   // TANK_CONTROL_6S.GTT_OUT_DATA.GTT_DemandsCompleted[2] := False;
   // TANK_CONTROL_6S.GTT_OUT_DATA.GTT_DemandsCompleted[1] := False;
   // TANK_CONTROL_6S.PVVX_OUT_DATA.PVVB_Alarms[14] := False;
   // TANK_CONTROL_6S.PVVX_OUT_DATA.PVVB_Alarms[13] := False;
   // TANK_CONTROL_6S.PVVX_OUT_DATA.PVVB_Alarms[12] := False;
   // TANK_CONTROL_6S.PVVX_OUT_DATA.PVVB_Alarms[11] := False;
   // TANK_CONTROL_6S.PVVX_OUT_DATA.PVVB_Alarms[10] := False;
   // TANK_CONTROL_6S.PVVX_OUT_DATA.PVVB_Alarms[9] := False;
   // TANK_CONTROL_6S.PVVX_OUT_DATA.PVVB_Alarms[8] := False;
   // TANK_CONTROL_6S.PVVX_OUT_DATA.PVVB_Alarms[7] := False;
   // TANK_CONTROL_6S.PVVX_OUT_DATA.PVVB_Alarms[6] := False;
   // TANK_CONTROL_6S.PVVX_OUT_DATA.PVVB_Alarms[5] := False;
   // TANK_CONTROL_6S.PVVX_OUT_DATA.PVVB_Alarms[4] := False;
   // TANK_CONTROL_6S.PVVX_OUT_DATA.PVVB_Alarms[3] := False;
   // TANK_CONTROL_6S.PVVX_OUT_DATA.PVVB_Alarms[2] := False;
   // TANK_CONTROL_6S.PVVX_OUT_DATA.PVVB_Alarms[1] := False;
   // TANK_CONTROL_6S.PVVX_OUT_DATA.PVVB_DemandsCompleted[14] := False;
   // TANK_CONTROL_6S.PVVX_OUT_DATA.PVVB_DemandsCompleted[13] := False;
   // TANK_CONTROL_6S.PVVX_OUT_DATA.PVVB_DemandsCompleted[12] := False;
   // TANK_CONTROL_6S.PVVX_OUT_DATA.PVVB_DemandsCompleted[11] := False;
   // TANK_CONTROL_6S.PVVX_OUT_DATA.PVVB_DemandsCompleted[10] := False;
   // TANK_CONTROL_6S.PVVX_OUT_DATA.PVVB_DemandsCompleted[9] := False;
   // TANK_CONTROL_6S.PVVX_OUT_DATA.PVVB_DemandsCompleted[8] := False;
   // TANK_CONTROL_6S.PVVX_OUT_DATA.PVVB_DemandsCompleted[7] := False;
   // TANK_CONTROL_6S.PVVX_OUT_DATA.PVVB_DemandsCompleted[6] := False;
   // TANK_CONTROL_6S.PVVX_OUT_DATA.PVVB_DemandsCompleted[5] := False;
   // TANK_CONTROL_6S.PVVX_OUT_DATA.PVVB_DemandsCompleted[4] := False;
   // TANK_CONTROL_6S.PVVX_OUT_DATA.PVVB_DemandsCompleted[3] := False;
   // TANK_CONTROL_6S.PVVX_OUT_DATA.PVVB_DemandsCompleted[2] := False;
   // TANK_CONTROL_6S.PVVX_OUT_DATA.PVVB_DemandsCompleted[1] := False;
   // TANK_CONTROL_6S.PVVX_OUT_DATA.PVVA_Alarms[14] := False;
   // TANK_CONTROL_6S.PVVX_OUT_DATA.PVVA_Alarms[13] := False;
   // TANK_CONTROL_6S.PVVX_OUT_DATA.PVVA_Alarms[12] := False;
   // TANK_CONTROL_6S.PVVX_OUT_DATA.PVVA_Alarms[11] := False;
   // TANK_CONTROL_6S.PVVX_OUT_DATA.PVVA_Alarms[10] := False;
   // TANK_CONTROL_6S.PVVX_OUT_DATA.PVVA_Alarms[9] := False;
   // TANK_CONTROL_6S.PVVX_OUT_DATA.PVVA_Alarms[8] := False;
   // TANK_CONTROL_6S.PVVX_OUT_DATA.PVVA_Alarms[7] := False;
   // TANK_CONTROL_6S.PVVX_OUT_DATA.PVVA_Alarms[6] := False;
   // TANK_CONTROL_6S.PVVX_OUT_DATA.PVVA_Alarms[5] := False;
   // TANK_CONTROL_6S.PVVX_OUT_DATA.PVVA_Alarms[4] := False;
   // TANK_CONTROL_6S.PVVX_OUT_DATA.PVVA_Alarms[3] := False;
   // TANK_CONTROL_1P.DWELL_TIMER.IN := False;
   // TANK_CONTROL_1P.MONITOR_TIMER.IN := False;
   // TANK_CONTROL_1P.ReOx_InitialTargetpHLevelAchieved := False;
   // TANK_CONTROL_6S.PVVX_OUT_DATA.PVVA_Alarms[2] := False;
   // TANK_CONTROL_6S.PVVX_OUT_DATA.PVVA_Alarms[1] := False;
   // TANK_CONTROL_6S.PVVX_OUT_DATA.PVVA_DemandsCompleted[14] := False;
   // TANK_CONTROL_6S.PVVX_OUT_DATA.PVVA_DemandsCompleted[13] := False;
   // TANK_CONTROL_6S.PVVX_OUT_DATA.PVVA_DemandsCompleted[12] := False;
   // TANK_CONTROL_6S.PVVX_OUT_DATA.PVVA_DemandsCompleted[11] := False;
   // TANK_CONTROL_6S.PVVX_OUT_DATA.PVVA_DemandsCompleted[10] := False;
   // TANK_CONTROL_6S.PVVX_OUT_DATA.PVVA_DemandsCompleted[9] := False;
   // TANK_CONTROL_6S.PVVX_OUT_DATA.PVVA_DemandsCompleted[8] := False;
   // TANK_CONTROL_6S.PVVX_OUT_DATA.PVVA_DemandsCompleted[7] := False;
   // TANK_CONTROL_6S.PVVX_OUT_DATA.PVVA_DemandsCompleted[6] := False;
   // TANK_CONTROL_6S.PVVX_OUT_DATA.PVVA_DemandsCompleted[5] := False;
   // TANK_CONTROL_6S.PVVX_OUT_DATA.PVVA_DemandsCompleted[4] := False;
   // TANK_CONTROL_6S.PVVX_OUT_DATA.PVVA_DemandsCompleted[3] := False;
   // TANK_CONTROL_6S.PVVX_OUT_DATA.PVVA_DemandsCompleted[2] := False;
   // TANK_CONTROL_6S.PVVX_OUT_DATA.PVVA_DemandsCompleted[1] := False;
   // TANK_CONTROL_1P.TankIPData.TANK_GROUP_SPARE_DI_5 := False;
   // TANK_CONTROL_1P.TankIPData.TANK_GROUP_SPARE_DI_6 := False;
   // TANK_CONTROL_1P.TankIPData.TANK_GROUP_SPARE_DI_7 := False;
   // TANK_CONTROL_1P.TankIPData.GTT_ISOL_VALVE_OPEN := False;
   // TANK_CONTROL_1P.TankIPData.GTT_ISOL_VALVE_CLSD := False;
   // TANK_CONTROL_1P.TankIPData.BWT_LEVEL_HIHI := False;
   // TANK_CONTROL_1P.TankIPData.TANK_ALARM := False;
   // TANK_CONTROL_1P.TankIPData.SPARE_DI_7 := False;
   // TANK_CONTROL_1S.TankIPData.TANKS_PRESS_HIHI := False;
   // TANK_CONTROL_1S.TankIPData.TANK_GROUP_SPARE_DI_2 := False;
   // TANK_CONTROL_1S.TankIPData.TANK_GROUP_SPARE_DI_3 := False;
   // TANK_CONTROL_1S.TankIPData.TANK_GROUP_SPARE_DI_4 := False;
   // TANK_CONTROL_1S.TankIPData.TANK_GROUP_SPARE_DI_5 := False;
   // TANK_CONTROL_1S.TankIPData.TANK_GROUP_SPARE_DI_6 := False;
   // TANK_CONTROL_1S.TankIPData.TANK_GROUP_SPARE_DI_7 := False;
   // TANK_CONTROL_1S.TankIPData.GTT_ISOL_VALVE_OPEN := False;
   // TANK_CONTROL_6P.GTT_OUT_DATA.GTT_Alarms[14] := False;
   // TANK_CONTROL_6P.GTT_OUT_DATA.GTT_Alarms[13] := False;
   // TANK_CONTROL_6P.GTT_OUT_DATA.GTT_Alarms[12] := False;
   // TANK_CONTROL_6P.GTT_OUT_DATA.GTT_Alarms[11] := False;
   // TANK_CONTROL_6P.GTT_OUT_DATA.GTT_Alarms[10] := False;
   // TANK_CONTROL_6P.GTT_OUT_DATA.GTT_Alarms[9] := False;
   // TANK_CONTROL_6P.GTT_OUT_DATA.GTT_Alarms[8] := False;
   // TANK_CONTROL_6P.GTT_OUT_DATA.GTT_Alarms[7] := False;
   // TANK_CONTROL_6P.GTT_OUT_DATA.GTT_Alarms[6] := False;
   // TANK_CONTROL_6P.GTT_OUT_DATA.GTT_Alarms[5] := False;
   // TANK_CONTROL_6P.GTT_OUT_DATA.GTT_Alarms[4] := False;
   // TANK_CONTROL_6P.GTT_OUT_DATA.GTT_Alarms[3] := False;
   // TANK_CONTROL_6P.GTT_OUT_DATA.GTT_Alarms[2] := False;
   // TANK_CONTROL_6P.GTT_OUT_DATA.GTT_Alarms[1] := False;
   // TANK_CONTROL_6P.GTT_OUT_DATA.GTT_DemandsCompleted[14] := False;
   // TANK_CONTROL_6P.GTT_OUT_DATA.GTT_DemandsCompleted[13] := False;
   // TANK_CONTROL_6P.GTT_OUT_DATA.GTT_DemandsCompleted[12] := False;
   // TANK_CONTROL_6P.GTT_OUT_DATA.GTT_DemandsCompleted[11] := False;
   // TANK_CONTROL_6P.GTT_OUT_DATA.GTT_DemandsCompleted[10] := False;
   // TANK_CONTROL_6P.GTT_OUT_DATA.GTT_DemandsCompleted[9] := False;
   // TANK_CONTROL_6P.GTT_OUT_DATA.GTT_DemandsCompleted[8] := False;
   // TANK_CONTROL_6P.GTT_OUT_DATA.GTT_DemandsCompleted[7] := False;
   // TANK_CONTROL_6P.GTT_OUT_DATA.GTT_DemandsCompleted[6] := False;
   // TANK_CONTROL_6P.GTT_OUT_DATA.GTT_DemandsCompleted[5] := False;
   // TANK_CONTROL_6P.GTT_OUT_DATA.GTT_DemandsCompleted[4] := False;
   // TANK_CONTROL_6P.GTT_OUT_DATA.GTT_DemandsCompleted[3] := False;
   // TANK_CONTROL_6P.GTT_OUT_DATA.GTT_DemandsCompleted[2] := False;
   // TANK_CONTROL_6P.GTT_OUT_DATA.GTT_DemandsCompleted[1] := False;
   // TANK_CONTROL_6P.PVVX_OUT_DATA.PVVB_Alarms[14] := False;
   // TANK_CONTROL_6P.PVVX_OUT_DATA.PVVB_Alarms[13] := False;
   // TANK_CONTROL_6P.PVVX_OUT_DATA.PVVB_Alarms[12] := False;
   // TANK_CONTROL_6P.PVVX_OUT_DATA.PVVB_Alarms[11] := False;
   // TANK_CONTROL_6P.PVVX_OUT_DATA.PVVB_Alarms[10] := False;
   // TANK_CONTROL_6P.PVVX_OUT_DATA.PVVB_Alarms[9] := False;
   // TANK_CONTROL_6P.PVVX_OUT_DATA.PVVB_Alarms[8] := False;
   // TANK_CONTROL_6P.PVVX_OUT_DATA.PVVB_Alarms[7] := False;
   // TANK_CONTROL_6P.PVVX_OUT_DATA.PVVB_Alarms[6] := False;
   // TANK_CONTROL_6P.PVVX_OUT_DATA.PVVB_Alarms[5] := False;
   // TANK_CONTROL_6P.PVVX_OUT_DATA.PVVB_Alarms[4] := False;
   // TANK_CONTROL_6P.PVVX_OUT_DATA.PVVB_Alarms[3] := False;
   // TANK_CONTROL_6P.PVVX_OUT_DATA.PVVB_Alarms[2] := False;
   // TANK_CONTROL_6P.PVVX_OUT_DATA.PVVB_Alarms[1] := False;
   // TANK_CONTROL_6P.PVVX_OUT_DATA.PVVB_DemandsCompleted[14] := False;
   // TANK_CONTROL_6P.PVVX_OUT_DATA.PVVB_DemandsCompleted[13] := False;
   // TANK_CONTROL_6P.PVVX_OUT_DATA.PVVB_DemandsCompleted[12] := False;
   // TANK_CONTROL_6P.PVVX_OUT_DATA.PVVB_DemandsCompleted[11] := False;
   // TANK_CONTROL_6P.PVVX_OUT_DATA.PVVB_DemandsCompleted[10] := False;
   // TANK_CONTROL_6P.PVVX_OUT_DATA.PVVB_DemandsCompleted[9] := False;
   // TANK_CONTROL_6P.PVVX_OUT_DATA.PVVB_DemandsCompleted[8] := False;
   // TANK_CONTROL_6P.PVVX_OUT_DATA.PVVB_DemandsCompleted[7] := False;
   // TANK_CONTROL_6P.PVVX_OUT_DATA.PVVB_DemandsCompleted[6] := False;
   // TANK_CONTROL_6P.PVVX_OUT_DATA.PVVB_DemandsCompleted[5] := False;
   // TANK_CONTROL_1S.DWELL_TIMER.IN := False;
   // TANK_CONTROL_1S.MONITOR_TIMER.IN := False;
   // TANK_CONTROL_1S.ReOx_InitialTargetpHLevelAchieved := False;
   // TANK_CONTROL_6P.PVVX_OUT_DATA.PVVB_DemandsCompleted[4] := False;
   // TANK_CONTROL_6P.PVVX_OUT_DATA.PVVB_DemandsCompleted[3] := False;
   // TANK_CONTROL_6P.PVVX_OUT_DATA.PVVB_DemandsCompleted[2] := False;
   // TANK_CONTROL_6P.PVVX_OUT_DATA.PVVB_DemandsCompleted[1] := False;
   // TANK_CONTROL_6P.PVVX_OUT_DATA.PVVA_Alarms[14] := False;
   // TANK_CONTROL_6P.PVVX_OUT_DATA.PVVA_Alarms[13] := False;
   // TANK_CONTROL_6P.PVVX_OUT_DATA.PVVA_Alarms[12] := False;
   // TANK_CONTROL_6P.PVVX_OUT_DATA.PVVA_Alarms[11] := False;
   // TANK_CONTROL_6P.PVVX_OUT_DATA.PVVA_Alarms[10] := False;
   // TANK_CONTROL_6P.PVVX_OUT_DATA.PVVA_Alarms[9] := False;
   // TANK_CONTROL_6P.PVVX_OUT_DATA.PVVA_Alarms[8] := False;
   // TANK_CONTROL_6P.PVVX_OUT_DATA.PVVA_Alarms[7] := False;
   // TANK_CONTROL_6P.PVVX_OUT_DATA.PVVA_Alarms[6] := False;
   // TANK_CONTROL_6P.PVVX_OUT_DATA.PVVA_Alarms[5] := False;
   // TANK_CONTROL_6P.PVVX_OUT_DATA.PVVA_Alarms[4] := False;
   // TANK_CONTROL_6P.PVVX_OUT_DATA.PVVA_Alarms[3] := False;
   // TANK_CONTROL_6P.PVVX_OUT_DATA.PVVA_Alarms[2] := False;
   // TANK_CONTROL_6P.PVVX_OUT_DATA.PVVA_Alarms[1] := False;
   // TANK_CONTROL_6P.PVVX_OUT_DATA.PVVA_DemandsCompleted[14] := False;
   // TANK_CONTROL_6P.PVVX_OUT_DATA.PVVA_DemandsCompleted[13] := False;
   // TANK_CONTROL_6P.PVVX_OUT_DATA.PVVA_DemandsCompleted[12] := False;
   // TANK_CONTROL_6P.PVVX_OUT_DATA.PVVA_DemandsCompleted[11] := False;
   // TANK_CONTROL_6P.PVVX_OUT_DATA.PVVA_DemandsCompleted[10] := False;
   // TANK_CONTROL_6P.PVVX_OUT_DATA.PVVA_DemandsCompleted[9] := False;
   // TANK_CONTROL_6P.PVVX_OUT_DATA.PVVA_DemandsCompleted[8] := False;
   // TANK_CONTROL_6P.PVVX_OUT_DATA.PVVA_DemandsCompleted[7] := False;
   // TANK_CONTROL_6P.PVVX_OUT_DATA.PVVA_DemandsCompleted[6] := False;
   // TANK_CONTROL_6P.PVVX_OUT_DATA.PVVA_DemandsCompleted[5] := False;
   // TANK_CONTROL_6P.PVVX_OUT_DATA.PVVA_DemandsCompleted[4] := False;
   // TANK_CONTROL_6P.PVVX_OUT_DATA.PVVA_DemandsCompleted[3] := False;
   // TANK_CONTROL_6P.PVVX_OUT_DATA.PVVA_DemandsCompleted[2] := False;
   // TANK_CONTROL_6P.PVVX_OUT_DATA.PVVA_DemandsCompleted[1] := False;
   // TANK_CONTROL_1S.TankIPData.GTT_ISOL_VALVE_CLSD := False;
   // TANK_CONTROL_1S.TankIPData.BWT_LEVEL_HIHI := False;
   // TANK_CONTROL_1S.TankIPData.TANK_ALARM := False;
   // TANK_CONTROL_1S.TankIPData.SPARE_DI_7 := False;
   // TANK_CONTROL_2P.TankIPData.TANKS_PRESS_HIHI := False;
   // TANK_CONTROL_2P.TankIPData.TANK_GROUP_SPARE_DI_2 := False;
   // TANK_CONTROL_2P.TankIPData.TANK_GROUP_SPARE_DI_3 := False;
   // TANK_CONTROL_2P.TankIPData.TANK_GROUP_SPARE_DI_4 := False;
   // TANK_CONTROL_2P.TankIPData.TANK_GROUP_SPARE_DI_5 := False;
   // TANK_CONTROL_2P.TankIPData.TANK_GROUP_SPARE_DI_6 := False;
   // TANK_CONTROL_2P.TankIPData.TANK_GROUP_SPARE_DI_7 := False;
   // TANK_CONTROL_2P.TankIPData.GTT_ISOL_VALVE_OPEN := False;
   // TANK_CONTROL_2P.TankIPData.GTT_ISOL_VALVE_CLSD := False;
   // TANK_CONTROL_2P.TankIPData.BWT_LEVEL_HIHI := False;
   // TANK_CONTROL_2P.TankIPData.TANK_ALARM := False;
   // TANK_CONTROL_2P.TankIPData.SPARE_DI_7 := False;
   // TANK_CONTROL_5S.GTT_OUT_DATA.GTT_Alarms[14] := False;
   // TANK_CONTROL_5S.GTT_OUT_DATA.GTT_Alarms[13] := False;
   // TANK_CONTROL_5S.GTT_OUT_DATA.GTT_Alarms[12] := False;
   // TANK_CONTROL_5S.GTT_OUT_DATA.GTT_Alarms[11] := False;
   // TANK_CONTROL_5S.GTT_OUT_DATA.GTT_Alarms[10] := False;
   // TANK_CONTROL_5S.GTT_OUT_DATA.GTT_Alarms[9] := False;
   // TANK_CONTROL_5S.GTT_OUT_DATA.GTT_Alarms[8] := False;
   // TANK_CONTROL_5S.GTT_OUT_DATA.GTT_Alarms[7] := False;
   // TANK_CONTROL_5S.GTT_OUT_DATA.GTT_Alarms[6] := False;
   // TANK_CONTROL_5S.GTT_OUT_DATA.GTT_Alarms[5] := False;
   // TANK_CONTROL_5S.GTT_OUT_DATA.GTT_Alarms[4] := False;
   // TANK_CONTROL_5S.GTT_OUT_DATA.GTT_Alarms[3] := False;
   // TANK_CONTROL_5S.GTT_OUT_DATA.GTT_Alarms[2] := False;
   // TANK_CONTROL_5S.GTT_OUT_DATA.GTT_Alarms[1] := False;
   // TANK_CONTROL_5S.GTT_OUT_DATA.GTT_DemandsCompleted[14] := False;
   // TANK_CONTROL_5S.GTT_OUT_DATA.GTT_DemandsCompleted[13] := False;
   // TANK_CONTROL_5S.GTT_OUT_DATA.GTT_DemandsCompleted[12] := False;
   // TANK_CONTROL_5S.GTT_OUT_DATA.GTT_DemandsCompleted[11] := False;
   // TANK_CONTROL_5S.GTT_OUT_DATA.GTT_DemandsCompleted[10] := False;
   // TANK_CONTROL_5S.GTT_OUT_DATA.GTT_DemandsCompleted[9] := False;
   // TANK_CONTROL_5S.GTT_OUT_DATA.GTT_DemandsCompleted[8] := False;
   // TANK_CONTROL_5S.GTT_OUT_DATA.GTT_DemandsCompleted[7] := False;
   // TANK_CONTROL_5S.GTT_OUT_DATA.GTT_DemandsCompleted[6] := False;
   // TANK_CONTROL_5S.GTT_OUT_DATA.GTT_DemandsCompleted[5] := False;
   // TANK_CONTROL_5S.GTT_OUT_DATA.GTT_DemandsCompleted[4] := False;
   // TANK_CONTROL_5S.GTT_OUT_DATA.GTT_DemandsCompleted[3] := False;
   // TANK_CONTROL_5S.GTT_OUT_DATA.GTT_DemandsCompleted[2] := False;
   // TANK_CONTROL_5S.GTT_OUT_DATA.GTT_DemandsCompleted[1] := False;
   // TANK_CONTROL_5S.PVVX_OUT_DATA.PVVB_Alarms[14] := False;
   // TANK_CONTROL_5S.PVVX_OUT_DATA.PVVB_Alarms[13] := False;
   // TANK_CONTROL_5S.PVVX_OUT_DATA.PVVB_Alarms[12] := False;
   // TANK_CONTROL_5S.PVVX_OUT_DATA.PVVB_Alarms[11] := False;
   // TANK_CONTROL_5S.PVVX_OUT_DATA.PVVB_Alarms[10] := False;
   // TANK_CONTROL_5S.PVVX_OUT_DATA.PVVB_Alarms[9] := False;
   // TANK_CONTROL_5S.PVVX_OUT_DATA.PVVB_Alarms[8] := False;
   // TANK_CONTROL_5S.PVVX_OUT_DATA.PVVB_Alarms[7] := False;
   // TANK_CONTROL_5S.PVVX_OUT_DATA.PVVB_Alarms[6] := False;
   // TANK_CONTROL_5S.PVVX_OUT_DATA.PVVB_Alarms[5] := False;
   // TANK_CONTROL_5S.PVVX_OUT_DATA.PVVB_Alarms[4] := False;
   // TANK_CONTROL_5S.PVVX_OUT_DATA.PVVB_Alarms[3] := False;
   // TANK_CONTROL_5S.PVVX_OUT_DATA.PVVB_Alarms[2] := False;
   // TANK_CONTROL_5S.PVVX_OUT_DATA.PVVB_Alarms[1] := False;
   // TANK_CONTROL_5S.PVVX_OUT_DATA.PVVB_DemandsCompleted[14] := False;
   // TANK_CONTROL_5S.PVVX_OUT_DATA.PVVB_DemandsCompleted[13] := False;
   // TANK_CONTROL_2P.DWELL_TIMER.IN := False;
   // TANK_CONTROL_2P.MONITOR_TIMER.IN := False;
   // TANK_CONTROL_2P.ReOx_InitialTargetpHLevelAchieved := False;
   // TANK_CONTROL_5S.PVVX_OUT_DATA.PVVB_DemandsCompleted[12] := False;
   // TANK_CONTROL_5S.PVVX_OUT_DATA.PVVB_DemandsCompleted[11] := False;
   // TANK_CONTROL_5S.PVVX_OUT_DATA.PVVB_DemandsCompleted[10] := False;
   // TANK_CONTROL_5S.PVVX_OUT_DATA.PVVB_DemandsCompleted[9] := False;
   // TANK_CONTROL_5S.PVVX_OUT_DATA.PVVB_DemandsCompleted[8] := False;
   // TANK_CONTROL_5S.PVVX_OUT_DATA.PVVB_DemandsCompleted[7] := False;
   // TANK_CONTROL_5S.PVVX_OUT_DATA.PVVB_DemandsCompleted[6] := False;
   // TANK_CONTROL_5S.PVVX_OUT_DATA.PVVB_DemandsCompleted[5] := False;
   // TANK_CONTROL_5S.PVVX_OUT_DATA.PVVB_DemandsCompleted[4] := False;
   // TANK_CONTROL_5S.PVVX_OUT_DATA.PVVB_DemandsCompleted[3] := False;
   // TANK_CONTROL_5S.PVVX_OUT_DATA.PVVB_DemandsCompleted[2] := False;
   // TANK_CONTROL_5S.PVVX_OUT_DATA.PVVB_DemandsCompleted[1] := False;
   // TANK_CONTROL_5S.PVVX_OUT_DATA.PVVA_Alarms[14] := False;
   // TANK_CONTROL_5S.PVVX_OUT_DATA.PVVA_Alarms[13] := False;
   // TANK_CONTROL_5S.PVVX_OUT_DATA.PVVA_Alarms[12] := False;
   // TANK_CONTROL_5S.PVVX_OUT_DATA.PVVA_Alarms[11] := False;
   // TANK_CONTROL_5S.PVVX_OUT_DATA.PVVA_Alarms[10] := False;
   // TANK_CONTROL_5S.PVVX_OUT_DATA.PVVA_Alarms[9] := False;
   // TANK_CONTROL_5S.PVVX_OUT_DATA.PVVA_Alarms[8] := False;
   // TANK_CONTROL_5S.PVVX_OUT_DATA.PVVA_Alarms[7] := False;
   // TANK_CONTROL_5S.PVVX_OUT_DATA.PVVA_Alarms[6] := False;
   // TANK_CONTROL_5S.PVVX_OUT_DATA.PVVA_Alarms[5] := False;
   // TANK_CONTROL_5S.PVVX_OUT_DATA.PVVA_Alarms[4] := False;
   // TANK_CONTROL_5S.PVVX_OUT_DATA.PVVA_Alarms[3] := False;
   // TANK_CONTROL_5S.PVVX_OUT_DATA.PVVA_Alarms[2] := False;
   // TANK_CONTROL_5S.PVVX_OUT_DATA.PVVA_Alarms[1] := False;
   // TANK_CONTROL_5S.PVVX_OUT_DATA.PVVA_DemandsCompleted[14] := False;
   // TANK_CONTROL_5S.PVVX_OUT_DATA.PVVA_DemandsCompleted[13] := False;
   // TANK_CONTROL_5S.PVVX_OUT_DATA.PVVA_DemandsCompleted[12] := False;
   // TANK_CONTROL_5S.PVVX_OUT_DATA.PVVA_DemandsCompleted[11] := False;
   // TANK_CONTROL_5S.PVVX_OUT_DATA.PVVA_DemandsCompleted[10] := False;
   // TANK_CONTROL_5S.PVVX_OUT_DATA.PVVA_DemandsCompleted[9] := False;
   // TANK_CONTROL_5S.PVVX_OUT_DATA.PVVA_DemandsCompleted[8] := False;
   // TANK_CONTROL_5S.PVVX_OUT_DATA.PVVA_DemandsCompleted[7] := False;
   // TANK_CONTROL_5S.PVVX_OUT_DATA.PVVA_DemandsCompleted[6] := False;
   // TANK_CONTROL_5S.PVVX_OUT_DATA.PVVA_DemandsCompleted[5] := False;
   // TANK_CONTROL_5S.PVVX_OUT_DATA.PVVA_DemandsCompleted[4] := False;
   // TANK_CONTROL_5S.PVVX_OUT_DATA.PVVA_DemandsCompleted[3] := False;
   // TANK_CONTROL_5S.PVVX_OUT_DATA.PVVA_DemandsCompleted[2] := False;
   // TANK_CONTROL_5S.PVVX_OUT_DATA.PVVA_DemandsCompleted[1] := False;
   // TANK_CONTROL_2S.TankIPData.TANKS_PRESS_HIHI := False;
   // TANK_CONTROL_2S.TankIPData.TANK_GROUP_SPARE_DI_2 := False;
   // TANK_CONTROL_2S.TankIPData.TANK_GROUP_SPARE_DI_3 := False;
   // TANK_CONTROL_2S.TankIPData.TANK_GROUP_SPARE_DI_4 := False;
   // TANK_CONTROL_2S.TankIPData.TANK_GROUP_SPARE_DI_5 := False;
   // TANK_CONTROL_2S.TankIPData.TANK_GROUP_SPARE_DI_6 := False;
   // TANK_CONTROL_2S.TankIPData.TANK_GROUP_SPARE_DI_7 := False;
   // TANK_CONTROL_2S.TankIPData.GTT_ISOL_VALVE_OPEN := False;
   // TANK_CONTROL_2S.TankIPData.GTT_ISOL_VALVE_CLSD := False;
   // TANK_CONTROL_2S.TankIPData.BWT_LEVEL_HIHI := False;
   // TANK_CONTROL_2S.TankIPData.TANK_ALARM := False;
   // TANK_CONTROL_2S.TankIPData.SPARE_DI_7 := False;
   // TANK_CONTROL_3P.TankIPData.TANKS_PRESS_HIHI := False;
   // TANK_CONTROL_3P.TankIPData.TANK_GROUP_SPARE_DI_2 := False;
   // TANK_CONTROL_3P.TankIPData.TANK_GROUP_SPARE_DI_3 := False;
   // TANK_CONTROL_3P.TankIPData.TANK_GROUP_SPARE_DI_4 := False;
   // TANK_CONTROL_5P.GTT_OUT_DATA.GTT_Alarms[14] := False;
   // TANK_CONTROL_5P.GTT_OUT_DATA.GTT_Alarms[13] := False;
   // TANK_CONTROL_5P.GTT_OUT_DATA.GTT_Alarms[12] := False;
   // TANK_CONTROL_5P.GTT_OUT_DATA.GTT_Alarms[11] := False;
   // TANK_CONTROL_5P.GTT_OUT_DATA.GTT_Alarms[10] := False;
   // TANK_CONTROL_5P.GTT_OUT_DATA.GTT_Alarms[9] := False;
   // TANK_CONTROL_5P.GTT_OUT_DATA.GTT_Alarms[8] := False;
   // TANK_CONTROL_5P.GTT_OUT_DATA.GTT_Alarms[7] := False;
   // TANK_CONTROL_5P.GTT_OUT_DATA.GTT_Alarms[6] := False;
   // TANK_CONTROL_5P.GTT_OUT_DATA.GTT_Alarms[5] := False;
   // TANK_CONTROL_5P.GTT_OUT_DATA.GTT_Alarms[4] := False;
   // TANK_CONTROL_5P.GTT_OUT_DATA.GTT_Alarms[3] := False;
   // TANK_CONTROL_5P.GTT_OUT_DATA.GTT_Alarms[2] := False;
   // TANK_CONTROL_5P.GTT_OUT_DATA.GTT_Alarms[1] := False;
   // TANK_CONTROL_5P.GTT_OUT_DATA.GTT_DemandsCompleted[14] := False;
   // TANK_CONTROL_5P.GTT_OUT_DATA.GTT_DemandsCompleted[13] := False;
   // TANK_CONTROL_5P.GTT_OUT_DATA.GTT_DemandsCompleted[12] := False;
   // TANK_CONTROL_5P.GTT_OUT_DATA.GTT_DemandsCompleted[11] := False;
   // TANK_CONTROL_5P.GTT_OUT_DATA.GTT_DemandsCompleted[10] := False;
   // TANK_CONTROL_5P.GTT_OUT_DATA.GTT_DemandsCompleted[9] := False;
   // TANK_CONTROL_5P.GTT_OUT_DATA.GTT_DemandsCompleted[8] := False;
   // TANK_CONTROL_5P.GTT_OUT_DATA.GTT_DemandsCompleted[7] := False;
   // TANK_CONTROL_5P.GTT_OUT_DATA.GTT_DemandsCompleted[6] := False;
   // TANK_CONTROL_5P.GTT_OUT_DATA.GTT_DemandsCompleted[5] := False;
   // TANK_CONTROL_5P.GTT_OUT_DATA.GTT_DemandsCompleted[4] := False;
   // TANK_CONTROL_5P.GTT_OUT_DATA.GTT_DemandsCompleted[3] := False;
   // TANK_CONTROL_5P.GTT_OUT_DATA.GTT_DemandsCompleted[2] := False;
   // TANK_CONTROL_5P.GTT_OUT_DATA.GTT_DemandsCompleted[1] := False;
   // TANK_CONTROL_5P.PVVX_OUT_DATA.PVVB_Alarms[14] := False;
   // TANK_CONTROL_5P.PVVX_OUT_DATA.PVVB_Alarms[13] := False;
   // TANK_CONTROL_5P.PVVX_OUT_DATA.PVVB_Alarms[12] := False;
   // TANK_CONTROL_5P.PVVX_OUT_DATA.PVVB_Alarms[11] := False;
   // TANK_CONTROL_5P.PVVX_OUT_DATA.PVVB_Alarms[10] := False;
   // TANK_CONTROL_5P.PVVX_OUT_DATA.PVVB_Alarms[9] := False;
   // TANK_CONTROL_5P.PVVX_OUT_DATA.PVVB_Alarms[8] := False;
   // TANK_CONTROL_5P.PVVX_OUT_DATA.PVVB_Alarms[7] := False;
   // TANK_CONTROL_5P.PVVX_OUT_DATA.PVVB_Alarms[6] := False;
   // TANK_CONTROL_5P.PVVX_OUT_DATA.PVVB_Alarms[5] := False;
   // TANK_CONTROL_5P.PVVX_OUT_DATA.PVVB_Alarms[4] := False;
   // TANK_CONTROL_5P.PVVX_OUT_DATA.PVVB_Alarms[3] := False;
   // TANK_CONTROL_5P.PVVX_OUT_DATA.PVVB_Alarms[2] := False;
   // TANK_CONTROL_5P.PVVX_OUT_DATA.PVVB_Alarms[1] := False;
   // TANK_CONTROL_5P.PVVX_OUT_DATA.PVVB_DemandsCompleted[14] := False;
   // TANK_CONTROL_5P.PVVX_OUT_DATA.PVVB_DemandsCompleted[13] := False;
   // TANK_CONTROL_2S.DWELL_TIMER.IN := False;
   // TANK_CONTROL_2S.MONITOR_TIMER.IN := False;
   // TANK_CONTROL_2S.ReOx_InitialTargetpHLevelAchieved := False;
   // TANK_CONTROL_5P.PVVX_OUT_DATA.PVVB_DemandsCompleted[12] := False;
   // TANK_CONTROL_5P.PVVX_OUT_DATA.PVVB_DemandsCompleted[11] := False;
   // TANK_CONTROL_5P.PVVX_OUT_DATA.PVVB_DemandsCompleted[10] := False;
   // TANK_CONTROL_5P.PVVX_OUT_DATA.PVVB_DemandsCompleted[9] := False;
   // TANK_CONTROL_5P.PVVX_OUT_DATA.PVVB_DemandsCompleted[8] := False;
   // TANK_CONTROL_5P.PVVX_OUT_DATA.PVVB_DemandsCompleted[7] := False;
   // TANK_CONTROL_5P.PVVX_OUT_DATA.PVVB_DemandsCompleted[6] := False;
   // TANK_CONTROL_5P.PVVX_OUT_DATA.PVVB_DemandsCompleted[5] := False;
   // TANK_CONTROL_5P.PVVX_OUT_DATA.PVVB_DemandsCompleted[4] := False;
   // TANK_CONTROL_5P.PVVX_OUT_DATA.PVVB_DemandsCompleted[3] := False;
   // TANK_CONTROL_5P.PVVX_OUT_DATA.PVVB_DemandsCompleted[2] := False;
   // TANK_CONTROL_5P.PVVX_OUT_DATA.PVVB_DemandsCompleted[1] := False;
   // TANK_CONTROL_5P.PVVX_OUT_DATA.PVVA_Alarms[14] := False;
   // TANK_CONTROL_5P.PVVX_OUT_DATA.PVVA_Alarms[13] := False;
   // TANK_CONTROL_5P.PVVX_OUT_DATA.PVVA_Alarms[12] := False;
   // TANK_CONTROL_5P.PVVX_OUT_DATA.PVVA_Alarms[11] := False;
   // TANK_CONTROL_5P.PVVX_OUT_DATA.PVVA_Alarms[10] := False;
   // TANK_CONTROL_5P.PVVX_OUT_DATA.PVVA_Alarms[9] := False;
   // TANK_CONTROL_5P.PVVX_OUT_DATA.PVVA_Alarms[8] := False;
   // TANK_CONTROL_5P.PVVX_OUT_DATA.PVVA_Alarms[7] := False;
   // TANK_CONTROL_5P.PVVX_OUT_DATA.PVVA_Alarms[6] := False;
   // TANK_CONTROL_5P.PVVX_OUT_DATA.PVVA_Alarms[5] := False;
   // TANK_CONTROL_5P.PVVX_OUT_DATA.PVVA_Alarms[4] := False;
   // TANK_CONTROL_5P.PVVX_OUT_DATA.PVVA_Alarms[3] := False;
   // TANK_CONTROL_5P.PVVX_OUT_DATA.PVVA_Alarms[2] := False;
   // TANK_CONTROL_5P.PVVX_OUT_DATA.PVVA_Alarms[1] := False;
   // TANK_CONTROL_5P.PVVX_OUT_DATA.PVVA_DemandsCompleted[14] := False;
   // TANK_CONTROL_5P.PVVX_OUT_DATA.PVVA_DemandsCompleted[13] := False;
   // TANK_CONTROL_5P.PVVX_OUT_DATA.PVVA_DemandsCompleted[12] := False;
   // TANK_CONTROL_5P.PVVX_OUT_DATA.PVVA_DemandsCompleted[11] := False;
   // TANK_CONTROL_5P.PVVX_OUT_DATA.PVVA_DemandsCompleted[10] := False;
   // TANK_CONTROL_5P.PVVX_OUT_DATA.PVVA_DemandsCompleted[9] := False;
   // TANK_CONTROL_5P.PVVX_OUT_DATA.PVVA_DemandsCompleted[8] := False;
   // TANK_CONTROL_5P.PVVX_OUT_DATA.PVVA_DemandsCompleted[7] := False;
   // TANK_CONTROL_5P.PVVX_OUT_DATA.PVVA_DemandsCompleted[6] := False;
   // TANK_CONTROL_5P.PVVX_OUT_DATA.PVVA_DemandsCompleted[5] := False;
   // TANK_CONTROL_5P.PVVX_OUT_DATA.PVVA_DemandsCompleted[4] := False;
   // TANK_CONTROL_5P.PVVX_OUT_DATA.PVVA_DemandsCompleted[3] := False;
   // TANK_CONTROL_5P.PVVX_OUT_DATA.PVVA_DemandsCompleted[2] := False;
   // TANK_CONTROL_5P.PVVX_OUT_DATA.PVVA_DemandsCompleted[1] := False;
   // TANK_CONTROL_3P.TankIPData.TANK_GROUP_SPARE_DI_5 := False;
   // TANK_CONTROL_3P.TankIPData.TANK_GROUP_SPARE_DI_6 := False;
   // TANK_CONTROL_3P.TankIPData.TANK_GROUP_SPARE_DI_7 := False;
   // TANK_CONTROL_3P.TankIPData.GTT_ISOL_VALVE_OPEN := False;
   // TANK_CONTROL_3P.TankIPData.GTT_ISOL_VALVE_CLSD := False;
   // TANK_CONTROL_3P.TankIPData.BWT_LEVEL_HIHI := False;
   // TANK_CONTROL_3P.TankIPData.TANK_ALARM := False;
   // TANK_CONTROL_3P.TankIPData.SPARE_DI_7 := False;
   // TANK_CONTROL_3S.TankIPData.TANKS_PRESS_HIHI := False;
   // TANK_CONTROL_3S.TankIPData.TANK_GROUP_SPARE_DI_2 := False;
   // TANK_CONTROL_3S.TankIPData.TANK_GROUP_SPARE_DI_3 := False;
   // TANK_CONTROL_3S.TankIPData.TANK_GROUP_SPARE_DI_4 := False;
   // TANK_CONTROL_3S.TankIPData.TANK_GROUP_SPARE_DI_5 := False;
   // TANK_CONTROL_3S.TankIPData.TANK_GROUP_SPARE_DI_6 := False;
   // TANK_CONTROL_3S.TankIPData.TANK_GROUP_SPARE_DI_7 := False;
   // TANK_CONTROL_3S.TankIPData.GTT_ISOL_VALVE_OPEN := False;
   // TANK_CONTROL_4S.GTT_OUT_DATA.GTT_Alarms[14] := False;
   // TANK_CONTROL_4S.GTT_OUT_DATA.GTT_Alarms[13] := False;
   // TANK_CONTROL_4S.GTT_OUT_DATA.GTT_Alarms[12] := False;
   // TANK_CONTROL_4S.GTT_OUT_DATA.GTT_Alarms[11] := False;
   // TANK_CONTROL_4S.GTT_OUT_DATA.GTT_Alarms[10] := False;
   // TANK_CONTROL_4S.GTT_OUT_DATA.GTT_Alarms[9] := False;
   // TANK_CONTROL_4S.GTT_OUT_DATA.GTT_Alarms[8] := False;
   // TANK_CONTROL_4S.GTT_OUT_DATA.GTT_Alarms[7] := False;
   // TANK_CONTROL_4S.GTT_OUT_DATA.GTT_Alarms[6] := False;
   // TANK_CONTROL_4S.GTT_OUT_DATA.GTT_Alarms[5] := False;
   // TANK_CONTROL_4S.GTT_OUT_DATA.GTT_Alarms[4] := False;
   // TANK_CONTROL_4S.GTT_OUT_DATA.GTT_Alarms[3] := False;
   // TANK_CONTROL_4S.GTT_OUT_DATA.GTT_Alarms[2] := False;
   // TANK_CONTROL_4S.GTT_OUT_DATA.GTT_Alarms[1] := False;
   // TANK_CONTROL_4S.GTT_OUT_DATA.GTT_DemandsCompleted[14] := False;
   // TANK_CONTROL_4S.GTT_OUT_DATA.GTT_DemandsCompleted[13] := False;
   // TANK_CONTROL_4S.GTT_OUT_DATA.GTT_DemandsCompleted[12] := False;
   // TANK_CONTROL_4S.GTT_OUT_DATA.GTT_DemandsCompleted[11] := False;
   // TANK_CONTROL_4S.GTT_OUT_DATA.GTT_DemandsCompleted[10] := False;
   // TANK_CONTROL_4S.GTT_OUT_DATA.GTT_DemandsCompleted[9] := False;
   // TANK_CONTROL_4S.GTT_OUT_DATA.GTT_DemandsCompleted[8] := False;
   // TANK_CONTROL_4S.GTT_OUT_DATA.GTT_DemandsCompleted[7] := False;
   // TANK_CONTROL_4S.GTT_OUT_DATA.GTT_DemandsCompleted[6] := False;
   // TANK_CONTROL_4S.GTT_OUT_DATA.GTT_DemandsCompleted[5] := False;
   // TANK_CONTROL_4S.GTT_OUT_DATA.GTT_DemandsCompleted[4] := False;
   // TANK_CONTROL_4S.GTT_OUT_DATA.GTT_DemandsCompleted[3] := False;
   // TANK_CONTROL_4S.GTT_OUT_DATA.GTT_DemandsCompleted[2] := False;
   // TANK_CONTROL_4S.GTT_OUT_DATA.GTT_DemandsCompleted[1] := False;
   // TANK_CONTROL_4S.PVVX_OUT_DATA.PVVB_Alarms[14] := False;
   // TANK_CONTROL_4S.PVVX_OUT_DATA.PVVB_Alarms[13] := False;
   // TANK_CONTROL_4S.PVVX_OUT_DATA.PVVB_Alarms[12] := False;
   // TANK_CONTROL_4S.PVVX_OUT_DATA.PVVB_Alarms[11] := False;
   // TANK_CONTROL_4S.PVVX_OUT_DATA.PVVB_Alarms[10] := False;
   // TANK_CONTROL_4S.PVVX_OUT_DATA.PVVB_Alarms[9] := False;
   // TANK_CONTROL_4S.PVVX_OUT_DATA.PVVB_Alarms[8] := False;
   // TANK_CONTROL_4S.PVVX_OUT_DATA.PVVB_Alarms[7] := False;
   // TANK_CONTROL_4S.PVVX_OUT_DATA.PVVB_Alarms[6] := False;
   // TANK_CONTROL_4S.PVVX_OUT_DATA.PVVB_Alarms[5] := False;
   // TANK_CONTROL_4S.PVVX_OUT_DATA.PVVB_Alarms[4] := False;
   // TANK_CONTROL_4S.PVVX_OUT_DATA.PVVB_Alarms[3] := False;
   // TANK_CONTROL_4S.PVVX_OUT_DATA.PVVB_Alarms[2] := False;
   // TANK_CONTROL_4S.PVVX_OUT_DATA.PVVB_Alarms[1] := False;
   // TANK_CONTROL_4S.PVVX_OUT_DATA.PVVB_DemandsCompleted[14] := False;
   // TANK_CONTROL_4S.PVVX_OUT_DATA.PVVB_DemandsCompleted[13] := False;
   // TANK_CONTROL_3P.DWELL_TIMER.IN := False;
   // TANK_CONTROL_3P.MONITOR_TIMER.IN := False;
   // TANK_CONTROL_3P.ReOx_InitialTargetpHLevelAchieved := False;
   // TANK_CONTROL_4S.PVVX_OUT_DATA.PVVB_DemandsCompleted[12] := False;
   // TANK_CONTROL_4S.PVVX_OUT_DATA.PVVB_DemandsCompleted[11] := False;
   // TANK_CONTROL_4S.PVVX_OUT_DATA.PVVB_DemandsCompleted[10] := False;
   // TANK_CONTROL_4S.PVVX_OUT_DATA.PVVB_DemandsCompleted[9] := False;
   // TANK_CONTROL_4S.PVVX_OUT_DATA.PVVB_DemandsCompleted[8] := False;
   // TANK_CONTROL_4S.PVVX_OUT_DATA.PVVB_DemandsCompleted[7] := False;
   // TANK_CONTROL_4S.PVVX_OUT_DATA.PVVB_DemandsCompleted[6] := False;
   // TANK_CONTROL_4S.PVVX_OUT_DATA.PVVB_DemandsCompleted[5] := False;
   // TANK_CONTROL_4S.PVVX_OUT_DATA.PVVB_DemandsCompleted[4] := False;
   // TANK_CONTROL_4S.PVVX_OUT_DATA.PVVB_DemandsCompleted[3] := False;
   // TANK_CONTROL_4S.PVVX_OUT_DATA.PVVB_DemandsCompleted[2] := False;
   // TANK_CONTROL_4S.PVVX_OUT_DATA.PVVB_DemandsCompleted[1] := False;
   // TANK_CONTROL_4S.PVVX_OUT_DATA.PVVA_Alarms[14] := False;
   // TANK_CONTROL_4S.PVVX_OUT_DATA.PVVA_Alarms[13] := False;
   // TANK_CONTROL_4S.PVVX_OUT_DATA.PVVA_Alarms[12] := False;
   // TANK_CONTROL_4S.PVVX_OUT_DATA.PVVA_Alarms[11] := False;
   // TANK_CONTROL_4S.PVVX_OUT_DATA.PVVA_Alarms[10] := False;
   // TANK_CONTROL_4S.PVVX_OUT_DATA.PVVA_Alarms[9] := False;
   // TANK_CONTROL_4S.PVVX_OUT_DATA.PVVA_Alarms[8] := False;
   // TANK_CONTROL_4S.PVVX_OUT_DATA.PVVA_Alarms[7] := False;
   // TANK_CONTROL_4S.PVVX_OUT_DATA.PVVA_Alarms[6] := False;
   // TANK_CONTROL_4S.PVVX_OUT_DATA.PVVA_Alarms[5] := False;
   // TANK_CONTROL_4S.PVVX_OUT_DATA.PVVA_Alarms[4] := False;
   // TANK_CONTROL_4S.PVVX_OUT_DATA.PVVA_Alarms[3] := False;
   // TANK_CONTROL_4S.PVVX_OUT_DATA.PVVA_Alarms[2] := False;
   // TANK_CONTROL_4S.PVVX_OUT_DATA.PVVA_Alarms[1] := False;
   // TANK_CONTROL_4S.PVVX_OUT_DATA.PVVA_DemandsCompleted[14] := False;
   // TANK_CONTROL_4S.PVVX_OUT_DATA.PVVA_DemandsCompleted[13] := False;
   // TANK_CONTROL_4S.PVVX_OUT_DATA.PVVA_DemandsCompleted[12] := False;
   // TANK_CONTROL_4S.PVVX_OUT_DATA.PVVA_DemandsCompleted[11] := False;
   // TANK_CONTROL_4S.PVVX_OUT_DATA.PVVA_DemandsCompleted[10] := False;
   // TANK_CONTROL_4S.PVVX_OUT_DATA.PVVA_DemandsCompleted[9] := False;
   // TANK_CONTROL_4S.PVVX_OUT_DATA.PVVA_DemandsCompleted[8] := False;
   // TANK_CONTROL_4S.PVVX_OUT_DATA.PVVA_DemandsCompleted[7] := False;
   // TANK_CONTROL_4S.PVVX_OUT_DATA.PVVA_DemandsCompleted[6] := False;
   // TANK_CONTROL_4S.PVVX_OUT_DATA.PVVA_DemandsCompleted[5] := False;
   // TANK_CONTROL_4S.PVVX_OUT_DATA.PVVA_DemandsCompleted[4] := False;
   // TANK_CONTROL_4S.PVVX_OUT_DATA.PVVA_DemandsCompleted[3] := False;
   // TANK_CONTROL_4S.PVVX_OUT_DATA.PVVA_DemandsCompleted[2] := False;
   // TANK_CONTROL_4S.PVVX_OUT_DATA.PVVA_DemandsCompleted[1] := False;
   // TANK_CONTROL_3S.TankIPData.GTT_ISOL_VALVE_CLSD := False;
   // TANK_CONTROL_3S.TankIPData.BWT_LEVEL_HIHI := False;
   // TANK_CONTROL_3S.TankIPData.TANK_ALARM := False;
   // TANK_CONTROL_3S.TankIPData.SPARE_DI_7 := False;
   // TANK_CONTROL_4P.TankIPData.TANKS_PRESS_HIHI := False;
   // TANK_CONTROL_4P.TankIPData.TANK_GROUP_SPARE_DI_2 := False;
   // TANK_CONTROL_4P.TankIPData.TANK_GROUP_SPARE_DI_3 := False;
   // TANK_CONTROL_4P.TankIPData.TANK_GROUP_SPARE_DI_4 := False;
   // TANK_CONTROL_4P.TankIPData.TANK_GROUP_SPARE_DI_5 := False;
   // TANK_CONTROL_4P.TankIPData.TANK_GROUP_SPARE_DI_6 := False;
   // TANK_CONTROL_4P.TankIPData.TANK_GROUP_SPARE_DI_7 := False;
   // TANK_CONTROL_4P.TankIPData.GTT_ISOL_VALVE_OPEN := False;
   // TANK_CONTROL_4P.TankIPData.GTT_ISOL_VALVE_CLSD := False;
   // TANK_CONTROL_4P.TankIPData.BWT_LEVEL_HIHI := False;
   // TANK_CONTROL_4P.TankIPData.TANK_ALARM := False;
   // TANK_CONTROL_4P.TankIPData.SPARE_DI_7 := False;
   // TANK_CONTROL_4P.GTT_OUT_DATA.GTT_Alarms[14] := False;
   // TANK_CONTROL_4P.GTT_OUT_DATA.GTT_Alarms[13] := False;
   // TANK_CONTROL_4P.GTT_OUT_DATA.GTT_Alarms[12] := False;
   // TANK_CONTROL_4P.GTT_OUT_DATA.GTT_Alarms[11] := False;
   // TANK_CONTROL_4P.GTT_OUT_DATA.GTT_Alarms[10] := False;
   // TANK_CONTROL_4P.GTT_OUT_DATA.GTT_Alarms[9] := False;
   // TANK_CONTROL_4P.GTT_OUT_DATA.GTT_Alarms[8] := False;
   // TANK_CONTROL_4P.GTT_OUT_DATA.GTT_Alarms[7] := False;
   // TANK_CONTROL_4P.GTT_OUT_DATA.GTT_Alarms[6] := False;
   // TANK_CONTROL_4P.GTT_OUT_DATA.GTT_Alarms[5] := False;
   // TANK_CONTROL_4P.GTT_OUT_DATA.GTT_Alarms[4] := False;
   // TANK_CONTROL_4P.GTT_OUT_DATA.GTT_Alarms[3] := False;
   // TANK_CONTROL_4P.GTT_OUT_DATA.GTT_Alarms[2] := False;
   // TANK_CONTROL_4P.GTT_OUT_DATA.GTT_Alarms[1] := False;
   // TANK_CONTROL_4P.GTT_OUT_DATA.GTT_DemandsCompleted[14] := False;
   // TANK_CONTROL_4P.GTT_OUT_DATA.GTT_DemandsCompleted[13] := False;
   // TANK_CONTROL_4P.GTT_OUT_DATA.GTT_DemandsCompleted[12] := False;
   // TANK_CONTROL_4P.GTT_OUT_DATA.GTT_DemandsCompleted[11] := False;
   // TANK_CONTROL_4P.GTT_OUT_DATA.GTT_DemandsCompleted[10] := False;
   // TANK_CONTROL_4P.GTT_OUT_DATA.GTT_DemandsCompleted[9] := False;
   // TANK_CONTROL_4P.GTT_OUT_DATA.GTT_DemandsCompleted[8] := False;
   // TANK_CONTROL_4P.GTT_OUT_DATA.GTT_DemandsCompleted[7] := False;
   // TANK_CONTROL_4P.GTT_OUT_DATA.GTT_DemandsCompleted[6] := False;
   // TANK_CONTROL_4P.GTT_OUT_DATA.GTT_DemandsCompleted[5] := False;
   // TANK_CONTROL_4P.GTT_OUT_DATA.GTT_DemandsCompleted[4] := False;
